(* Logix 5000 project; controller PLC_MCC1300_75F1 vendor 1 type 14 code 166 rev 32.11; software revision 32.04; part 9 of 83 *)

        [36].xFaulted := 1, [36].dEntryStatus := 16#0000_3000, [36].dFaultCode := 16#0000_0204, [36].dInstance := 16#0000_2268, [37].xConnected := 1, [37].xFaulted := 1, [37].dEntryStatus := 16#0000_3000, [37].dFaultCode := 16#0000_0204, [37].dInstance := 16#0000_494b, [38].xConnected := 1, [38].xFaulted := 1, [38].dEntryStatus := 16#0000_3000, [38].dFaultCode := 16#0000_0204, [38].dInstance := 16#0000_de82, [39].xConnected := 1, [39].xFaulted := 1, [39].dEntryStatus := 16#0000_3000, [39].dFaultCode := 16#0000_0204, [39].dInstance := 16#0000_ad3d, [40].xConnected := 1, [40].xFaulted := 1, [40].dEntryStatus := 16#0000_3000, [40].dFaultCode := 16#0000_0204, [40].dInstance := 16#0000_11ec, [41].xFaulted := 1, [41].dEntryStatus := 16#0000_1000, [41].dFaultCode := 16#0000_0204, [41].dInstance := 16#0000_7d3f, [42].xConnected := 1, [42].xFaulted := 1, [42].dEntryStatus := 16#0000_3000, [42].dFaultCode := 16#0000_0204, [42].dInstance := 16#0000_cb26, [43].xConnected := 1, [43].xFaulted := 1, [43].dEntryStatus := 16#0000_3000, [43].dFaultCode := 16#0000_0204, [43].dInstance := 16#0000_9dd1, [44].xConnected := 1, [44].xFaulted := 1, [44].dEntryStatus := 16#0000_3000, [44].dFaultCode := 16#0000_0204, [44].dInstance := 16#0000_2cb0, [45].xConnected := 1, [45].xFaulted := 1, [45].dEntryStatus := 16#0000_3000, [45].dFaultCode := 16#0000_0204, [45].dInstance := 16#0000_3773, [46].xConnected := 1, [46].xFaulted := 1, [46].dEntryStatus := 16#0000_3000, [46].dFaultCode := 16#0000_0204, [46].dInstance := 16#0000_0d0a, [47].xConnected := 1, [47].dEntryStatus := 16#0000_4000, [47].dInstance := 16#0000_f22b, [48].xConnected := 1, [48].dEntryStatus := 16#0000_4000, [48].dInstance := 16#0000_f6c7, [49].xConnected := 1,
        [49].dEntryStatus := 16#0000_4000, [49].dInstance := 16#0000_de7a); {access Read Only}
        [0]   // ETH_MCC1300
        [11]   // M3AZ01
        [12]   // M3AZ02
        [13]   // M3AZ03
        [14]   // M3AZ04
        [15]   // M3AZ05
        [16]   // M3AZ06
        [17]   // M3AZ07
        [18]   // M3AZ08
        [72]   // E93AZ1
        [31]   // TDKAZ05N
        [32]   // TDKAZ05S
        [33]   // TDAZ00N
        [34]   // TDAZ00S
        [35]   // TDAZ01N
        [36]   // TDAZ01S
        [37]   // TDAZ02N
        [19]   // M3AZ09
        [73]   // E96AZ1
        [75]   // E98AZ1
        [74]   // E97AZ1
        [20]   // M3AZ10
        [21]   // TDKAZ00N
        [38]   // TDAZ02S
        [39]   // TDAZ03N
        [40]   // TDAZ03S
        [41]   // TDAZ04N
        [42]   // TDAZ04S
        [43]   // TDAZ05N
        [44]   // TDAZ05S
        [50]   // E53AZ1
        [46]   // D010M1PM1
        [47]   // D010M2PM1
        [61]   // E77AZ1
        [62]   // E78AZ1
        [48]   // D020PM1
        [51]   // E61AZ1
        [52]   // E62AZ1
        [63]   // E81AZ1
        [64]   // E82AZ1
        [54]   // E64AZ1
        [53]   // E63AZ1
        [55]   // E65AZ1
        [65]   // E83AZ1
        [66]   // E84AZ1
        [56]   // E66AZ1
        [57]   // E67AZ1
        [58]   // E71AZ1
        [67]   // E85AZ1
        [68]   // E86AZ1
        [5]   // TD5680AP1
        [59]   // E73AZ1
        [60]   // E76AZ1
        [69]   // E87AZ1
        [70]   // E88AZ1
        [71]   // E91AZ1
        [1]   // ETH_M2
        [6]   // M3683AP1
        [7]   // E152AP1
        [8]   // RIOM13
        [22]   // TDKAZ00S
        [23]   // TDKAZ01N
        [24]   // TDKAZ01S
        [25]   // TDKAZ02N
        [26]   // TDKAZ02S
        [27]   // TDKAZ03N
        [28]   // TDKAZ03S
        [29]   // TDKAZ04N
        [30]   // TDKAZ04S
   MMI_DATA : INT[64] := ([1] := 4088, [2] := 4095, [8] := 4095, [11] := 2048, [20] := -1, [21] := -1, [22] := 1, [23] := 1);   // MMI DATA For Fix 32
        [12].0   // FIX MMI VMCC M2 Panel Overtemp Alarm
        [12].1   // FIX MMI VMCC TD Panel Overtemp Alarm
   MMI_FROM_MB : MESSAGE;
        MessageParameters(ServiceCode := 16#004b, LocalElement := MMI_DATA[20], ...)
   MMI_TO_MB : MESSAGE;
        MessageParameters(ServiceCode := 16#004c, LocalElement := MMI_DATA[0], ...)
   MMI_TO_MB_N15 : MESSAGE;
        MessageParameters(ServiceCode := 16#004c, LocalElement := MMI_DATA[0], ...)
   MS_LEHR : ALIAS FOR N20[11];
   MS_LINE : ALIAS FOR N20[13];
   MS_TRIM : ALIAS FOR N20[12];
   N10 : DINT[50] := ([10] := 2100, [40] := 4095);
        [16].1   // LEHR SPEED Speed received From Reliance Capping system is Valid
        [16].0   // LEHR SPEED Speed received From Reliance AutoMax PLC Is Valid
   N100 : DINT[1];
   N105 : DINT[1];
   N11 : DINT[500];
        [96]   // VISION INTERFACE: 2ND MOST CURRNET REJECTION REASON
        [97]   // VISION INTERFACE: 3RD MOST CURRNET REJECTION REASON
        [94].1   // Host & HMI Read Data: No Data From Vision System
        [94].2   // Host & HMI Read Data: Not Used Reserved for Focus CPS
        [94].3   // Host & HMI Read Data: Not Used Reserved for Focus CPS
        [94].4   // Host & HMI Read Data: Not Used Reserved for Focus CPS
        [79]   // Powder Camera Inspected Plate host IDENT
        [80]   // Host & HMI Read Data: Vision Broken Plate Count
        [81]   // Host & HMI Read Data: Vision Width Error Count
        [82]   // Host & HMI Read Data: Vision Length Error Count
        [83]   // Host & HMI Read Data: Vision Edge Defect Count
        [84]   // Host & HMI Read Data: Vision Corner Defect Count
        [85]   // Host & HMI Read Data: Vision Skew Count
        [86]   // Host & HMI Read Data: Vision Squareness Count
        [87]   // Host & HMI Read Data: Vision Fault Mark Count
        [88]   // Host & HMI Read Data: Vision Plate Missing Count
        [89]   // Host & HMI Read Data: Vision Not Separated Count
        [90]   // Host & HMI Read Data: Vision Other Count
        [91]   // Host & HMI Read Data: Vision Good Pieces Count
        [94].7   // Host & HMI Read Data: Vision System Is Disabled
        [92]   // Host & HMI Read Data: Vision Bad Pieces Count
        [93]   // Host & HMI Read Data: Vision No Response Count
        [94]   // Host & HMI Read Data: Vision Status Word
        [95]   // VISION INTERFACE: MOST CURRNET REJECTION REASON
        [94].0   // Host & HMI Read Data: All Pieces Are Bad
        [94].5   // Host & HMI Read Data: Vision System Is Online
        [94].6   // Host & HMI Read Data: Vision Service Required
   N110 : DINT[1];
   N115 : DINT[1];
   N11_HOST : INT[500] := ([0] := 22347, [1] := 22347, [20] := 9447, [21] := 96, [22] := 2047, [23] := 2047, [24] := 21845, [25] := 21, [26] := 53, [27] := 53, [38] := 2, [40] := 1, [60] := 554, [61] := 13, [62] := 20, [63] := 528, [65] := 609, [66] := 576, [67] := 4736, [68] := 453, [69] := 4902, [70] := 1028, [72] := 1536, [73] := 8320, [74] := 1, [79] := 8320, [80] := 1, [94] := 1, [101] := 648, [102] := 3, [103] := 204, [104] := 22347, [131] := 647, [133] := 45, [134] := 22346, [141] := 646, [143] := 45, [144] := 22346); {produced}
   N12 : DINT[500];
        [0]   // When this is Non-zero host Computer has Written new
        [3]   // HOST WRITE DATA: Glass Thickness (mils)
        [5]   // HOST WRITE DATA: Packing Station In Use Bits
        [6]   // HOST WRITE DATA: Ribbon Type (32=Eclipse Adv)
        [60]   // New cap data Buffer written by Host Computer
   N120 : DINT[1];
   N125 : DINT[1];
   N12_HOST : INT[500] := ([0] := 1, [1] := 650, [2] := 233, [3] := 15, [4] := 7653, [6] := 32, [7] := 31); {produced}
   N13 : DINT[500];
   N130 : INT[8] := ([0] := 1, [1] := 1, [2] := 1, [4] := 1325, [5] := 1, [6] := 1, [7] := 1);
        [3].10   // M2 -->> M4 Reliance Handoff Sensor (Redundant - on South side)
        [5].0   // M2-->M4 Benchboard No. 1 crusher Down
        [5].1   // M2-->M4 Benchboard No. 1 crusher Pushbutton
        [3].14   // M2 -->> M4 Crush all Selector Switch
        [3].15   // M2 -->> M4 Re-allocate To crusher Push-button
        [3].12   // M2 -->> M4 SPARE
        [3].1   // M2 -->> M4 SPARE
        [3].11   // M2 -->> M4
        [3].13   // M2 -->> M4 SPARE
        [3].2   // M2 -->> M4 SPARE
        [3].3   // M2 -->> M4 SPARE
        [3].4   // M2 -->> M4 SPARE
        [3].5   // M2 -->> M4 SPARE
        [3].6   // M2 -->> M4 SPARE
        [3].7   // M2 -->> M4 SPARE
        [3].8   // M2 -->> M4 SPARE
        [3].9   // M2 -->> M4 SPARE
   N131 : INT[8] := ([1] := 132, [4] := 450);
        [3].9   // M4 -->> M2 Reject Window Lamp
        [1]   // M2 -->> M4 Copy mainline Crusher status bits from M2 to M4
        [5].0   // M4-->M2 Float Glass Prodution
        [5].1   // M4-->M2 UL Crusher Is Faulted
        [3].14   // M4 -->> M2 ML is in Sleep Mode
        [3].3   // M4 -->> M2 Mainline Sec. Trans. Drive Fault
        [3].5   // M4 -->> M2 Mainline Sec. Trans. E-Stop
        [3].6   // M4 -->> M2 Mainline Sec. Trans. Backup
        [5].2   // M4-->M2 VISION SYS Rejected Plate Alarm Horn
        [1].11   // M4 -->> M2 Mainline vision Conveyor Stopped
        [3].10   // M4 -->> M2 Leg 2 Is In Sleep Mode Transfer Unavailable
        [3].11   // M4 -->> M2 Leg 3 Is In Sleep Mode Transfer Unavailable
        [3].12   // M4 -->> M2 Leg 4 Is In Sleep Mode Transfer Unavailable
        [3].13   // M4 -->> M2 Leg 5 Is In Sleep Mode Transfer Unavailable
        [4]   // M4 -->> M2 Trim speed
        [3].8   // M4 -->> M2 Reliance Data Received
        [3].15   // M4 -->> M2 M4 Heartbeat
        [3].1   // M4 -->> M2 SPARE
        [3].2   // M4 -->> M2 SPARE
   N135 : DINT[10];
        [0].12   // VHSC BTW Error Bit
        [5].12   // VHSC BTR Error Bit
        [0].15   // VHSC BTW Enable Bit
        [5].15   // VHSC BTR Enable Bit
   N136 : DINT[64];
        [1].15   // VHSC Data Representation Mode 0 = Binary 1 = BCD
        [30].0   // Output 01 Output/Counter Mapping Bits PC00
        [30].1   // Output 01 Output/Counter Mapping Bits PC01
        [30].2   // Output 01 Output/Counter Mapping Bits PC02
        [30].3   // Output 01 Output/Counter Mapping Bits PC03
        [1].0   // Reset PC00 - ACTIVE HIGH !
        [25].0   // Output 00 Output/Counter Mapping Bits PC00
        [25].1   // Output 00 Output/Counter Mapping Bits PC01
        [25].2   // Output 00 Output/Counter Mapping Bits PC02
        [25].3   // Output 00 Output/Counter Mapping Bits PC03
        [25]   // *************** * Output 00 ** * Mapping ** * Bits ** ***************
        [1].1   // Reset PC01 - ACTIVE HIGH !
        [21]   // Counter 0 Sample Period X 10mS
        [22]   // Counter 1 Sample Period X 10mS
        [1].2   // Reset PC02 - ACTIVE HIGH !
        [3]   // Mode Bits For Counters 0 and 1 ** Default ** ** Used **
        [13]   // PC00 Preset Value MSD
        [1].8   // PC00 Load Preset-
        [1].9   // PC01 Load Preset-
        [14]   // PC00 Preset Value LSD
        [15]   // PC01 Preset Value MSD
        [1].4   // PC00 New Data Acknowledge
        [2].10   // Output 02 Force
        [26]   // Output 00 ON VALUE MSD
        [10]   // PC02 Rollover Value LSD
        [11]   // PC03 Rollover Value LSD
        [12]   // PC03 Rollover Value LSD
        [16]   // PC01 Preset Value LSD
        [17]   // PC02 Preset Value MSD
        [18]   // PC02 Preset Value LSD
        [19]   // PC03 Preset Value LSD
        [1].10   // PC02 Load Preset-
        [1].11   // PC03 Load Preset-
        [5]   // PC00 Rollover Value MSD
        [1]   // Word 1 VHSC BTW Data
        [1].3   // Reset PC03 - ACTIVE HIGH !
        [6]   // PC00 Rollover Value LSD
        [7]   // PC01 Rollover Value MSD
        [1].12   // Not Used
        [1].13   // Not Used
        [1].14   // Not Used
        [1].5   // PC01 New Data Acknowledge
        [1].6   // PC03 New Data Acknowledge
        [1].7   // PC02 New Data Acknowledge
        [2].11   // Output 03 Force
        [2].12   // Output 04 Force
        [23]   // Counter 2 Sample Period X 10mS
        [24]   // Counter 3 Sample Period X 10mS
        [30]   // *************** * Output 01 ** * Mapping ** * Bits ** ***************
        [27]   // Output 00 ON VALUE LSD
        [31]   // Output 01 ON VALUE MSD
        [28]   // Output 00 OFF VALUE MSD
        [29]   // Output 00 OFF VALUE LSD
        [2]   // Word 2 VHSC BTW Data
        [2].0   // Output 00 Enable
        [2].1   // Output 01 Enable
        [2].13   // Output 05 Force
        [2].14   // Output 06 Force
        [2].15   // Output 07 Force
        [2].2   // Output 02 Enable
        [2].3   // Output 03 Enable
        [2].4   // Output 04 Enable
        [2].5   // Output 05 Enable
        [2].6   // Output 06 Enable
        [2].7   // Output 07 Enable
        [2].8   // Output 00 Force
        [2].9   // Output 01 Force
        [35]   // *************** * Output 02 ** * Mapping ** * Bits ** ***************
        [32]   // Output 01 ON VALUE LSD
        [36]   // Output 02 ON VALUE MSD
        [33]   // Output 01 OFF VALUE MSD
        [34]   // Output 01 OFF VALUE LSD
        [40]   // *************** * Output 03 ** * Mapping ** * Bits ** ***************
        [37]   // Output 02 ON VALUE LSD
        [46]   // Output 04 ON VALUE MSD
        [38]   // Output 02 OFF VALUE MSD
        [39]   // Output 02 OFF VALUE LSD
        [45]   // *************** * Output 04 ** * Mapping ** * Bits ** ***************
        [50]   // *************** * Output 05 ** * Mapping ** * Bits ** ***************
        [47]   // Output 04 ON VALUE LSD
        [56]   // Output 06 ON VALUE MSD
        [48]   // Output 04 OFF VALUE MSD
        [49]   // Output 04 OFF VALUE LSD
        [55]   // *************** * Output 06 ** * Mapping ** * Bits ** ***************
        [60]   // *************** * Output 07 ** * Mapping ** * Bits ** ***************
        [57]   // Output 06 ON VALUE LSD
        [61]   // Output 07 ON VALUE MSD
        [58]   // Output 06 OFF VALUE MSD
        [59]   // Output 06 OFF VALUE LSD
        [8]   // PC01 Rollover Value LSD
        [62]   // Output 07 ON VALUE LSD
        [63]   // Output 07 OFF VALUE MSD
        [9]   // PC02 Rollover Value MSD
   N137 : DINT[18];
   N138 : DINT[18];
   N139 : DINT[18];
        [1].0   // Successful First BTW after program start
        [2].10   // VHSC-PC02 Gate Input
        [1]   // VHSC status word No.1
        [1].10   // VHSC Gate Input
        [1].11   // VHSC Gate Input
        [2].8   // VHSC-PC00 Gate Input
        [10]   // PC03 Count LSD
        [2]   // VHSC status word No.2
        [1].8   // VHSC Gate Input
        [1].9   // VHSC Gate Input
        [2].0   // OUTPUT 00 Status
        [2].1   // OUTPUT 01 Status
        [2].12   // VHSC-PC03
        [2].13   // not used
        [2].15   // not used
        [2].2   // OUTPUT 02 Status
        [2].3   // OUTPUT 03 Status
        [2].4   // OUTPUT 04 Status
        [2].5   // OUTPUT 05 Status
        [2].6   // OUTPUT 06 Status
        [2].7   // OUTPUT 07 Status
        [2].9   // VHSC-PC01 Gate Input
        [3]   // PC00 Count MSD
        [4]   // PC00 Count LSD
        [5]   // PC01 Count MSD
        [6]   // PC01 Count LSD
        [7]   // PC02 Count MSD
        [8]   // PC02 Count LSD
        [9]   // PC03 Count LSD
   N14 : DINT[500] := ([61] := 4088, [62] := 4095, [68] := 4095, [71] := 2048, [80] := -1, [81] := -1, [82] := 1, [83] := 1, [240] := 6, [250] := 3313, [251] := 782, [260] := 7, [460] := 1, [469] := 258, [470] := 1, [479] := 258, [480] := -1, [488] := 256, [489] := 256, [490] := -1, [496] := 256, [497] := 256, [498] := 256, [499] := 256);
        [252].10   // TRIM DECK Trim Zone 5 North knocker Move Up
        [252].11   // TRIM DECK Trim Zone 5 South knocker Move Up
        [250].10   // TRIM DECK Trim Zone 5 North trim Auto mode
        [251].10   // TRIM DECK Trim Zone 5 North trim Manual mode
        [255]   // TRIM KNOCKERS Remapped inputs for all Move out Selector Sws.
        [273]   // TRIM DECK NTH Out Sel. Sw. Examine Masked Move Result
        [272]   // TRIM DECK NTH In Sel. Sw. Examine Masked Move Result
        [61]   // HOST/MMI READ Word containing Bits for drive Fault NORTH
        [253].10   // TRIM DECK Trim Zone 5 North knocker Move Down
        [240].1   // Float Glass Hold Down Wheels Manual Raise
        [256].0   // TRIM DECK Krurl drop North deck Move In
        [275]   // TRIM DECK STH In Sel. Sw. Examine Masked Move Result
        [253].2   // TRIM DECK Trim Zone 1 North knocker Move Down
        [276]   // TRIM DECK STH Out Sel. Sw. Examine Masked Move Result
        [251].11   // TRIM DECK Trim Zone 5 South trim Manual mode
        [253].3   // TRIM DECK Trim Zone 1 South knocker Move Down
        [256].1   // TRIM DECK Krurl drop South deck Move In
        [240].0   // Float Glass Hold Down Wheels Automatic Mode
        [250].2   // TRIM DECK Trim Zone 1 North trim Auto mode
        [260].0   // TRIM KNOCKERS Permissive to Start adj drive 1 = Drive idle 0 = Drv in use
        [255].10   // TRIM DECK Trim Zone 5 North knocker Move Out
        [255].11   // TRIM DECK Trim Zone 5 South knocker Move Out
        [271]   // TRIM DECK NTH Contactor Examine Masked Move Result
        [274]   // TRIM DECK STH Contactor Examine Masked Move Result
        [68]   // HOST/MMI READ Word containing Foward bits For Conveyors
        [253].4   // TRIM DECK Trim Zone 2 North knocker Move Down
        [253].5   // TRIM DECK Trim Zone 2 South knocker Move Down
        [253].6   // TRIM DECK Trim Zone 3 North knocker Move Down
        [253].7   // TRIM DECK Trim Zone 3 South knocker Move Down
        [254]   // TRIM KNOCKERS Remapped inputs for all Move in Selector Sws.
        [251].0   // TRIM DECK Krurl drop North trim Manual mode
        [460]   // TD MMI Zone 4 South Skew Adjustment
        [240].3   // Eclipse Hold Down Wheels Manual Raise
        [90].0   // To Float 1 host, bars on/off
        [312]   // HMI Data: Transfer 1A Stopping Offset for Rotated Glass [in x 10]
        [302]   // HMI Data: Transfer 1 Stopping Offset for Rotated Glass [in x 10]
        [351]   // HMI Read & Write Data: Transfer 1 Take All Cap Length
        [253].8   // TRIM DECK Trim Zone 4 North knocker Move Down
        [240].2   // Eclipse Hold Down Wheels Auto Mode
        [253].9   // TRIM DECK Trim Zone 4 South knocker Move Down
        [250].11   // TRIM DECK Trim Zone 5 South trim Auto mode
        [253].11   // TRIM DECK Trim Zone 5 South knocker Move Down
        [62]   // HOST/MMI READ Word containing Bits for drive Fault SOUTH AND 1-3
        [72].0   // FIX MMI VMCC M2 Panel Overtemp Alarm
        [72].1   // FIX MMI VMCC TD Panel Overtemp Alarm
        [470]   // TD MMI Zone 5 South Skew Adjustment
        [480]   // TD MMI Zone 3 South Skew Adjustment
        [490]   // TD MMI Zone 2 South Skew Adjustment
        [250]   // TRIM DECK Word containing All auto mode Bits
        [62].0   // Host Read Conv 1 Fault
        [251].2   // TRIM DECK Trim Zone 1 North trim Manual mode
        [250].3   // TRIM DECK Trim Zone 1 South trim Auto mode
        [61].10   // Host Read Conv 11N Fault
        [251].3   // TRIM DECK Trim Zone 1 South trim Manual mode
        [251].4   // TRIM DECK Trim Zone 2 North trim Manual mode
        [251].5   // TRIM DECK Trim Zone 2 South trim Manual mode
        [62].1   // Host Read Conv 2 Fault
        [61].11   // Host Read Conv 12N Fault
        [254].10   // TRIM DECK Trim Zone 5 North knocker Move In
        [254].11   // TRIM DECK Trim Zone 5 South knocker Move In
        [251].6   // TRIM DECK Trim Zone 3 North trim Manual mode
        [256].2   // TRIM DECK Trim Zone 1 North deck Move In
        [250].0   // TRIM DECK Krurl drop North trim Auto mode
        [250].4   // TRIM DECK Trim Zone 2 North trim Auto mode
        [256].3   // TRIM DECK Trim Zone 1 South deck Move In
        [251].7   // TRIM DECK Trim Zone 3 South trim Manual mode
        [251].8   // TRIM DECK Trim Zone 4 North trim Manual mode
        [256].4   // TRIM DECK Trim Zone 2 North deck Move In
        [251].9   // TRIM DECK Trim Zone 4 South trim Manual mode
        [256].5   // TRIM DECK Trim Zone 2 South deck Move In
        [250].1   // TRIM DECK Krurl drop South trim Auto mode
        [250].5   // TRIM DECK Trim Zone 2 South trim Auto mode
        [256].6   // TRIM DECK Trim Zone 3 North deck Move In
        [253].0   // TRIM DECK Krurl drop North knocker Move Down
        [253].1   // TRIM DECK Krurl drop South knocker Move Down
        [255].2   // TRIM DECK Trim Zone 1 North knocker Move Out
        [255].3   // TRIM DECK Trim Zone 1 South knocker Move Out
        [255].4   // TRIM DECK Trim Zone 2 North knocker Move Out
        [255].5   // TRIM DECK Trim Zone 2 South knocker Move Out
        [255].6   // TRIM DECK Trim Zone 3 North knocker Move Out
        [255].7   // TRIM DECK Trim Zone 3 South knocker Move Out
        [255].8   // TRIM DECK Trim Zone 4 North knocker Move Out
        [255].9   // TRIM DECK Trim Zone 4 South knocker Move Out
        [257].2   // TRIM DECK Trim Zone 1 North deck Move Out
        [256].7   // TRIM DECK Trim Zone 3 South deck Move In
        [257].3   // TRIM DECK Trim Zone 1 South deck Move Out
        [256].8   // TRIM DECK Trim Zone 4 North deck Move In
        [250].6   // TRIM DECK Trim Zone 3 North trim Auto mode
        [250].7   // TRIM DECK Trim Zone 3 South trim Auto mode
        [250].8   // TRIM DECK Trim Zone 4 North trim Auto mode
        [256].9   // TRIM DECK Trim Zone 4 South deck Move In
        [257].0   // TRIM DECK Krurl drop North deck Move Out
        [251].1   // TRIM DECK Krurl drop South trim Manual mode
        [252].2   // TRIM DECK Trim Zone 1 North knocker Move Up
        [257].4   // TRIM DECK Trim Zone 2 North deck Move Out
        [252].3   // TRIM DECK Trim Zone 1 South knocker Move Up
        [252].4   // TRIM DECK Trim Zone 2 North knocker Move Up
        [252].5   // TRIM DECK Trim Zone 2 South knocker Move Up
        [252].6   // TRIM DECK Trim Zone 3 North knocker Move Up
        [252].7   // TRIM DECK Trim Zone 3 South knocker Move Up
        [250].9   // TRIM DECK Trim Zone 4 South trim Auto mode
        [252].0   // TRIM DECK Krurl drop North knocker Move Up
        [252].1   // TRIM DECK Krurl drop South knocker Move Up
        [254].0   // TRIM DECK Krurl drop North knocker Move In
        [254].1   // TRIM DECK Krurl drop South knocker Move In
        [256].10   // TRIM DECK Trim Zone 5 North deck Move In
        [256].11   // TRIM DECK Trim Zone 5 South deck Move In
        [252].8   // TRIM DECK Trim Zone 4 North knocker Move Up
        [252].9   // TRIM DECK Trim Zone 4 South knocker Move Up
        [254].2   // TRIM DECK Trim Zone 1 North knocker Move In
        [254].3   // TRIM DECK Trim Zone 1 South knocker Move In
        [254].4   // TRIM DECK Trim Zone 2 North knocker Move In
        [254].5   // TRIM DECK Trim Zone 2 South knocker Move In
        [254].6   // TRIM DECK Trim Zone 3 North knocker Move In
        [254].7   // TRIM DECK Trim Zone 3 South knocker Move In
        [254].8   // TRIM DECK Trim Zone 4 North knocker Move In
        [254].9   // TRIM DECK Trim Zone 4 South knocker Move In
        [255].0   // TRIM DECK Krurl drop North knocker Move Out
        [255].1   // TRIM DECK Krurl drop South knocker Move Out
        [257].10   // TRIM DECK Trim Zone 5 North deck Move Out
        [257].11   // TRIM DECK Trim Zone 5 South deck Move Out
        [257].1   // TRIM DECK Krurl drop South deck Move Out
        [62].2   // Host Read Conv 3 Fault
        [84]   // HMI Write Data: Vision Edge On Defect Tol. [mm x 10]
        [112]   // HMI Write Data: Vision -Skew Tolerance [deg x 100]
        [80]   // HMI Write Data: Vision Over Width Tolerance [mm x 10]
        [301]   // HMI Data: Transfer 1 TE Stopping Position [in x 10]
        [257].5   // TRIM DECK Trim Zone 2 South deck Move Out
        [61].9   // Host Read Conv 10N Fault
        [62].9   // Host Read Conv 10S Fault
        [61].3   // Host Read Conv 4N Fault
        [257].6   // TRIM DECK Trim Zone 3 North deck Move Out
        [81]   // HMI Write Data: Vision Over Length Tolerance [mm x 10]
        [85]   // HMI Write Data: Vision Corner On Defect Tol. [mm x 10]
        [311]   // HMI Data: Transfer 1A TE Stopping Position [in x 10]
        [257].7   // TRIM DECK Trim Zone 3 South deck Move Out
        [110]   // HMI Write Data: Vision Under Width Tolerance [mm x 10]
        [111]   // HMI Write Data: Vision Under Length Tolerance [mm x 10]
        [114]   // HMI Write Data: Vision Edge Off Defect Tol. [mm x 10]
        [115]   // HMI Write Data: Vision Corner Off Defect Tol. [mm x 10]
        [170]   // MMI 400 DECK OP Adjust Distance For Larger Plates [in]
        [257].8   // TRIM DECK Trim Zone 4 North deck Move Out
        [250].12   // TRIM DECK SPARE
        [250].13   // TRIM DECK SPARE
        [250].14   // TRIM DECK SPARE
        [250].15   // TRIM DECK SPARE
        [251].12   // TRIM DECK SPARE
        [251].13   // TRIM DECK SPARE
        [251].14   // TRIM DECK SPARE
        [251].15   // TRIM DECK SPARE
        [252].12   // TRIM DECK SPARE
        [252].13   // TRIM DECK SPARE
        [252].14   // TRIM DECK SPARE
        [252].15   // TRIM DECK SPARE
        [253].12   // TRIM DECK SPARE
        [253].13   // TRIM DECK SPARE
        [253].14   // TRIM DECK SPARE
        [253].15   // TRIM DECK SPARE
        [254].12   // TRIM DECK SPARE
        [254].13   // TRIM DECK SPARE
        [254].14   // TRIM DECK SPARE
        [254].15   // TRIM DECK SPARE
        [255].12   // TRIM DECK SPARE
        [255].13   // TRIM DECK SPARE
        [255].14   // TRIM DECK SPARE
        [255].15   // TRIM DECK SPARE
        [256].12   // TRIM DECK SPARE
        [256].13   // TRIM DECK SPARE
        [256].14   // TRIM DECK SPARE
        [256].15   // TRIM DECK SPARE
        [257].12   // TRIM DECK SPARE
        [257].13   // TRIM DECK SPARE
        [257].14   // TRIM DECK SPARE
        [257].15   // TRIM DECK SPARE
        [257].9   // TRIM DECK Trim Zone 4 South deck Move Out
        [260].1   // TRIM DECK NTH Permissive to Start adj drive 1 = Drive idle 0 = Drv in use
        [260].2   // TRIM DECK STH Permissive to Start adj drive 1 = Drive idle 0 = Drv in use
        [62].10   // Host Read Conv 11S Fault
        [62].11   // Host Read Conv 12S Fault
        [61].4   // Host Read Conv 5N Fault
        [61].5   // Host Read Conv 6N Fault
        [61].6   // Host Read Conv 7N Fault
        [61].7   // Host Read Conv 8N Fault
        [61].8   // Host Read Conv 9N Fault
        [62].3   // Host Read Conv 4S Fault
        [62].4   // Host Read Conv 5S Fault
        [62].5   // Host Read Conv 6S Fault
        [62].6   // Host Read Conv 7S Fault
        [62].7   // Host Read Conv 8S Fault
        [62].8   // Host Read Conv 9S Fault
        [113]   // HMI Write Data: Vision -Squareness Tol. [mm x 10]
        [350]   // HMI Read & Write Data: Transfer 1 Take All Cap ID
        [358]   // HMI Read & Write Data: Transfer 1 Size A Split Width
        [82]   // HMI Write Data: Vision +Skew Tolerance [deg x 100]
        [83]   // HMI Write Data: Vision +Squareness Tol. [mm x 10]
        [86]   // HMI Write Data: Glass Substrate Type
   N14_HOST : INT[999]; {produced}
   N15 : DINT[500];
   N16 : DINT[500];
   N17 : DINT[100];
   N177 : DINT[10] := ([0] := 56, [1] := 1, [2] := 80, [5] := 2);
   N178 : DINT[100];
   N179 : DINT[100];
   N18 : DINT[100];
   N184 : DINT[50] := ([0] := 13, [1] := 94, [2] := 95, [3] := 96, [4] := 97, [5] := 98, [6] := 99, [7] := 100, [8] := 101, [9] := 4096, [10] := 11, [11] := 911, [12] := 671, [14] := 695, [16] := 23, [17] := 47, [18] := 107, [20] := 4, [21] := 139, [22] := 140, [23] := 141, [24] := 142, [25] := 143, [26] := 144, [27] := 145, [28] := 146, [29] := 8, [30] := 2, [31] := 902, [32] := 798, [34] := 686, [37] := 109, [49] := 2048);
   N185 : DINT[1];
   N187 : DINT[1];
   N188 : DINT[48] := ([4] := 256, [6] := 3840, [8] := 1280, [10] := 1280, [12] := 1280, [14] := 1280, [16] := 1280, [18] := 1280, [20] := 3328, [22] := 3840, [24] := 3840, [26] := 3840, [28] := 3840, [30] := 256);
   N189 : DINT[40];
   N190 : DINT[40];
   N191 : DINT[64];
   N192 : DINT[40];
   N193 : DINT[40] := ([0] := -22773, [1] := -27996, [5] := 1, [6] := 98, [7] := 1, [8] := 1, [17] := 102, [18] := 1, [20] := 96, [21] := 96, [22] := 97, [23] := 96, [24] := 97, [25] := 6, [26] := 103, [27] := 98, [28] := 98, [29] := 99, [30] := 474, [31] := 393, [32] := 96, [33] := 380);
   N194 : DINT[45] := ([2] := 166, [3] := 419, [4] := 166, [5] := 213, [7] := 206, [14] := -26651, [15] := 25346, [16] := 18332, [17] := -17337, [18] := 424, [19] := 19629, [20] := 169, [21] := 13674, [27] := 8, [29] := 1, [37] := 8114, [39] := 11259, [41] := 5595);
   N195 : DINT[40] := ([0] := 26204, [1] := 26204, [5] := 3, [7] := 1);
   N196 : DINT[1];
   N197 : DINT[1];
   N198 : DINT[1];
   N199 : DINT[1];
   N20 : DINT[50] := ([1] := 200, [2] := 500, [3] := 1200, [4] := 3000, [11] := 600, [12] := 150, [13] := 67, [14] := 40);
        [12]   // Milliseconds for two inches of glass travel at TRIM SPEED
        [11]   // Milliseconds for 2 inches of glass travel at LEHR SPEED
        [13]   // Milliseconds for 2 inches of glass travel at LINE SPEED
        [4]   // Runout Speed
        [1]   // Lehr Speed
        [2]   // Trim Speed
        [3]   // Line-Speed
   N200 : DINT[160];
   N201 : DINT[100];
   N202 : DINT[100];
   N203 : DINT[100];
   N204 : DINT[100];
   N205 : DINT[100];
   N206 : DINT[100];
   N207 : DINT[100];
   N208 : DINT[100];
   N209 : DINT[100];
   N21 : DINT[31] := ([0] := 2, [1] := 6144, [2] := 8320, [14] := 128);
        [0].5   // PLC -->> Copro Force Baseline/ Threshold (Set by MMI and Reset on LE)
        [0].2   // PLC -->> Copro Send Test Message to Vision
        [0].8   // PLC -->> Copro Reset Request for Baseline (Pushbutton at Vision)
        [0].3   // PLC -->> Copro No Update (From MMI)
        [14].8   // Copro -->> PLC Sending Test Message
        [14].0   // Copro -->> PLC All Bad Msg From Vision (Flashing Red)
        [14].1   // Copro -->> PLC No Data Msg From Vision (Solid Red)
        [0].1   // New data is Ready for VISCOMM Cleared by MLVISION
        [3]   // VISCOM Result Register --------------- 1=Good! 2=BAD!
        [0].4   // PLC --> Copro Reset Vision Counters (From VAX)
        [14].4   // Copro -->> PLC Doing Baseline (Flashing Blue)
        [14].5   // Copro -->> PLC Doing Threshold (Flasing Blue)
        [3].1   // VISCOM Result Register --------------- 1=Good! 2=Bad!
        [14].7   // Copro -->> PLC Copro Request for Baseline (Solid Blue)
        [3].0   // VISCOM Result Register --------------- 1 = Good 2 = Bad!
        [0].14   // PLC -->> Copro Used by VISCOM
        [14].6   // Copro -->> PLC Waiting
        [14].14   // Copro -->> PLC Bad Checksum
        [14].15   // Copro -->> PLC Bad Response
        [1]   // VISCOM New Length data (64ths)
        [2]   // VISCOM New Width data (64ths)
        [0].0   // PLC -->> Copro Debug
   N210 : DINT[100];
   N211 : DINT[100];
   N212 : DINT[100];
   N213 : DINT[100];
   N214 : DINT[100];
   N214_1 : ALIAS FOR N214[1];
   N214_5 : ALIAS FOR N214[5];
   N215 : DINT[100];
   N216 : DINT[100];
   N217 : DINT[100];
   N218 : DINT[100];
   N219 : DINT[100];
   N220 : DINT[100];
   N221 : DINT[100];
   N222 : DINT[100];
   N223 : DINT[100];
   N224 : DINT[100];
   N225 : DINT[100];
   N226 : DINT[100];
   N227 : DINT[100];
   N228 : DINT[100];
   N229 : DINT[100];
   N230 : DINT[100];
   N231 : DINT[100];
   N232 : DINT[100];
   N25 : DINT[110] := ([0] := 774, [1] := 1, [2] := 1, [3] := 1, [4] := 1, [5] := 1, [100] := 774);
        [1].1   // Vision System Results Buffer: Service Required for Vision System
        [3]   // Vision System Results Buffer: Number of Streams across Conveyor
        [0]   // Vision System Results Buffer: Group ID
        [2]   // Vision System Results Buffer: New data Flag (1 = New data)
        [100]   // Vision System Results PLC ID DTR Change of Value Reference
        [10]   // Vision System Results Buffer: Split 2B Reject Flag
        [11]   // Vision System Results Buffer: Split 2C Reject Flag
        [12]   // Vision System Results Buffer: Split 2D Reject Flag
        [13]   // Vision System Results Buffer: Split 3A Reject Flag
        [14]   // Vision System Results Buffer: Split 3B Reject Flag
        [15]   // Vision System Results Buffer: Split 3C Reject Flag
        [16]   // Vision System Results Buffer: Split 3D Reject Flag
        [17]   // Vision System Results Buffer: Split 4A Reject Flag
        [18]   // Vision System Results Buffer: Split 4B Reject Flag
        [19]   // Vision System Results Buffer: Split 4C Reject Flag
        [20]   // Vision System Results Buffer: Split 4D Reject Flag
        [21]   // Vision System Results Buffer: Split 5A Reject Flag
        [22]   // Vision System Results Buffer: Split 5B Reject Flag
        [23]   // Vision System Results Buffer: Split 5C Reject Flag
        [24]   // Vision System Results Buffer: Split 5D Reject Flag
        [25]   // Vision System Results Buffer: Split 6A Reject Flag
        [5]   // Vision System Results Buffer: Split 1A Reject Flag
        [6]   // Vision System Results Buffer: Split 1B Reject Flag
        [7]   // Vision System Results Buffer: Split 1C Reject Flag
        [26]   // Vision System Results Buffer: Split 6B Reject Flag
        [27]   // Vision System Results Buffer: Split 6C Reject Flag
        [28]   // Vision System Results Buffer: Split 6D Reject Flag
        [29]   // Vision System Results Buffer: Split 7A Reject Flag
        [30]   // Vision System Results Buffer: Split 7B Reject Flag
        [31]   // Vision System Results Buffer: Split 7C Reject Flag
        [32]   // Vision System Results Buffer: Split 7D Reject Flag
        [33]   // Vision System Results Buffer: Split 8A Reject Flag
        [34]   // Vision System Results Buffer: Split 8B Reject Flag
        [35]   // Vision System Results Buffer: Split 8C Reject Flag
        [36]   // Vision System Results Buffer: Split 8D Reject Flag
        [37]   // Vision System Results Buffer: Split 9A Reject Flag
        [38]   // Vision System Results Buffer: Split 9B Reject Flag
        [39]   // Vision System Results Buffer: Split 9C Reject Flag
        [40]   // Vision System Results Buffer: Split 9D Reject Flag
        [8]   // Vision System Results Buffer: Split 1D Reject Flag
        [9]   // Vision System Results Buffer: Split 2A Reject Flag
        [1]   // Vision System Results Buffer: Eagle-I Status Word
        [1].0   // Vision System Results Buffer: Vision System is Online
        [4]   // Vision System Results Buffer: Number of Splits down Conveyor
   N26 : DINT[150] := ([0] := 774, [2] := 3123, [3] := 1, [4] := 1, [5] := 12, [6] := 12, [7] := 1500, [8] := 32, [9] := 24, [10] := 32, [11] := 12, [12] := 12, [13] := 1500, [14] := 32, [15] := 24, [16] := 56, [17] := 8320, [21] := 5062, [100] := 20480, [101] := 774, [102] := 512, [105] := -22762, [106] := 2378, [107] := 23012, [108] := 4404, [109] := 22405, [110] := 846, [111] := -32768);
        [100].10   // VISION INTFCE: Cap Detected Entering Vision is a GOOD Plate with NO Splits
        [100].12   // VISION INTERFACE: Ignore Length Measurements on Queued Plates
        [100].2   // VISION INTERFACE: Results for New Cap ID Are Detected
        [100].4   // VISION INTERFACE: Cap Entering Conv 14 Check for Vis Required
        [100].8   // VIS INTFCE: Inspected Cap Prim Destination is Leg 1 or Leg 1A or L3
        [102].2   // one shot for Leading Edge of Data Valid Signal from Vision Sys
        [102].3   // VISION INTFCE: Bit to Reset Vision Debug Counters (Manually set)
        [102].8   // One shot for Glass Type Changing to Eclipse Advantage
        [104].0   // VIS INTFCE: No Vis Results Received for Glass Passing Thru X1 toward 1A
        [104].1   // VIS INTFCE: Inspection Results Not Received AND Glass is being Thrown Away
        [105]   // VISION INTERFACE: DEBUG COUNTER # of Good Plates from Data Packet
        [106]   // VISION INTERFACE: DEBUG COUNTER # of Bad Plates from Data Packet
        [107]   // VISION INTERFACE: DEBUG COUNTER # of Uninspected Plates from Data
        [109]   // VISION INTERFACE: DEBUG COUNTER # of Bad Plates from I/O Signals
        [13]   // Vision System Input Datafile: Neg Skew Tolerance [deg x 100]
        [100].9   // VIS INTFCE: Inspected Cap is a Leg 2 ; 4; or 5 Cap
        [100].3   // VISION INTERFACE: OK to Use New Vision Results
        [102].9   // One shot for Glass Type Changing to Base Glass
        [17]   // Vision System Input Datafile: Stream A Width [64ths]
        [18]   // Vision System Input Datafile: Stream B Width [64ths]
        [19]   // Vision System Input Datafile: Stream C Width [64ths]
        [20]   // Vision System Input Datafile: Stream D Width [64ths]
        [21]   // Vision System Input Datafile: Split 1 Length [64ths]
        [22]   // Vision System Input Datafile: Split 2 Length [64ths]
        [30].0   // Vision System Input Datafile: Stream A Inspect bit for Split 1
        [30].1   // Vision System Input Datafile: Stream A Inspect bit for Split 2
        [30].2   // Vision System Input Datafile: Stream A Inspect bit for Split 3
        [30].3   // Vision System Input Datafile: Stream A Inspect bit for Split 4
        [30].4   // Vision System Input Datafile: Stream A Inspect bit for Split 5
        [30].5   // Vision System Input Datafile: Stream A Inspect bit for Split 6
        [30].6   // Vision System Input Datafile: Stream A Inspect bit for Split 7
        [30].7   // Vision System Input Datafile: Stream A Inspect bit for Split 8
        [30].8   // Vision System Input Datafile: Stream A Inspect bit for Split 9
        [31].0   // Vision System Input Datafile: Stream B Inspect bit for Split 1
        [31].1   // Vision System Input Datafile: Stream B Inspect bit for Split 2
        [31].2   // Vision System Input Datafile: Stream B Inspect bit for Split 3
        [31].3   // Vision System Input Datafile: Stream B Inspect bit for Split 4
        [31].4   // Vision System Input Datafile: Stream B Inspect bit for Split 5
        [31].5   // Vision System Input Datafile: Stream B Inspect bit for Split 6
        [31].6   // Vision System Input Datafile: Stream B Inspect bit for Split 7
        [31].7   // Vision System Input Datafile: Stream B Inspect bit for Split 8
        [31].8   // Vision System Input Datafile: Stream B Inspect bit for Split 9
        [32].0   // Vision System Input Datafile: Stream C Inspect bit for Split 1
        [32].1   // Vision System Input Datafile: Stream C Inspect bit for Split 2
        [32].2   // Vision System Input Datafile: Stream C Inspect bit for Split 3
        [32].3   // Vision System Input Datafile: Stream C Inspect bit for Split 4
        [32].4   // Vision System Input Datafile: Stream C Inspect bit for Split 5
        [32].5   // Vision System Input Datafile: Stream C Inspect bit for Split 6
        [32].6   // Vision System Input Datafile: Stream C Inspect bit for Split 7
        [32].7   // Vision System Input Datafile: Stream C Inspect bit for Split 8
        [32].8   // Vision System Input Datafile: Stream C Inspect bit for Split 9
        [33].0   // Vision System Input Datafile: Stream D Inspect bit for Split 1
        [33].1   // Vision System Input Datafile: Stream D Inspect bit for Split 2
        [33].2   // Vision System Input Datafile: Stream D Inspect bit for Split 3
        [33].3   // Vision System Input Datafile: Stream D Inspect bit for Split 4
        [33].4   // Vision System Input Datafile: Stream D Inspect bit for Split 5
        [33].5   // Vision System Input Datafile: Stream D Inspect bit for Split 6
        [33].6   // Vision System Input Datafile: Stream D Inspect bit for Split 7
        [33].7   // Vision System Input Datafile: Stream D Inspect bit for Split 8
        [33].8   // Vision System Input Datafile: Stream D Inspect bit for Split 9
        [100].7   // VISION INTERFACE: Piece Called Bad By Vision Sys
        [102].10   // One shot for Glass Type Changing to Mirrorpane
        [34]   // Vision System Input Datafile: Quality Code for Split 1
        [35]   // Vision System Input Datafile: Quality Code for Split 2
        [36]   // Vision System Input Datafile: Quality Code for Split 3
        [37]   // Vision System Input Datafile: Quality Code for Split 4
        [38]   // Vision System Input Datafile: Quality Code for Split 5
        [39]   // Vision System Input Datafile: Quality Code for Split 6
        [40]   // Vision System Input Datafile: Quality Code for Split 7
        [15]   // Vision System Input Datafile: Neg Edge Tolerance [64ths]
        [6]   // Vision System Input Datafile: Pos Length Tolerance [64ths]
        [41]   // Vision System Input Datafile: Quality Code for Split 8
        [8]   // Vision System Input Datafile: Pos Square Tolerance [64ths]
        [99].0   // VISION INTERFACE: Primary Dest Cap Entering: Leg 1AN
        [99].1   // VISION INTERFACE: Primary Dest Cap Entering: Leg 1AS
        [99].2   // VISION INTERFACE: Primary Dest Cap Entering: Leg 1BN
        [99].4   // VISION INTERFACE: Primary Dest Cap Entering: Leg 2A LES
        [3]   // Vision System Input Datafile: Number of Streams across Conveyor
        [99].5   // VISION INTERFACE: Primary Dest Cap Entering: Leg 2B Robot
        [42]   // Vision System Input Datafile: Quality Code for Split 9
        [99]   // VISION INTERFACE: Primary Dest Cap Entering Vision Sys
        [1]   // Vision System Input Datafile: Substrate Type
        [100].5   // VISION INTERFACE: Cap Needs Vision Res Check for Receipt
        [100].0   // VISION INTERFACE: Cap Detected Entering the Vision System
        [23]   // Vision System Input Datafile: Split 3 Length [64ths]
        [24]   // Vision System Input Datafile: Split 4 Length [64ths]
        [9]   // Vision System Input Datafile: Pos Edge Tolerance [64ths]
        [11]   // Vision System Input Datafile: Neg Width Tolerance [64ths]
        [25]   // Vision System Input Datafile: Split 5 Length [64ths]
        [99].6   // VISION INTERFACE: Primary Dest Cap Entering: Mainline LES
        [99].3   // VISION INTERFACE: Primary Dest Cap Entering: Leg 1BS
        [100].15   // VISION INTERFACE: is Mirrorpane
        [0]   // Vision System Input Datafile: Group ID
        [101]   // VISION INTERFACE: PLC ID of Cap Entering Vision Sys
        [100].14   // VISION INTERFACE: Glass Type is Base glass
        [102].1   // One Shot for Glass Entering Conveyor 14
        [104].2   // VISION INTERFACE: Glass Type is Solar E
        [26]   // Vision System Input Datafile: Split 6 Length [64ths]
        [27]   // Vision System Input Datafile: Split 7 Length [64ths]
        [104].4   // VISION INTERFACE: Glass Type is TEC
        [28]   // Vision System Input Datafile: Split 8 Length [64ths]
        [29]   // Vision System Input Datafile: Split 9 Length [64ths]
        [104].5   // VISION INTERFACE: Glass Type is MirrorView
        [100].11   // VIS INTFCE: Glass Inspection Is in Progress
        [100].13   // VISION INTERFACE: Glass Type is Eclipse Adv
        [102].11   // One shot for Glass Type Changing to Solar E
        [103]   // VISION INTERFACE: Inspected Cap Primary Dest Word
        [30]   // Vision System Input Datafile: Stream A Inspect Word
        [31]   // Vision System Input Datafile: Stream B Inspect Word
        [32]   // Vision System Input Datafile: Stream C Inspect Word
        [33]   // Vision System Input Datafile: Stream D Inspect Word
        [100].6   // VISION INTERFACE: Piece Called Good By Vision Sys
        [102].12   // One shot for Glass Type Changing to Blue Active
        [2]   // Vision System Input Datafile: Substrate Thickness [64ths]
        [104].3   // VISION INTERFACE: Glass Type is Blue Active
        [102].0   // One Shot for Glass Entering Vision System
        [5]   // Vision System Input Datafile: Pos Width Tolerance [64ths]
        [100].1   // VISION INTERFACE: New Data Copied from Vision Output
        [10]   // Vision System Input Datafile: Pos Corner Tolerance [64ths]
        [12]   // Vision System Input Datafile: Neg Length Tolerance [64ths]
        [14]   // Vision System Input Datafile: Neg Square Tolerance [64ths]
        [16]   // Vision System Input Datafile: Neg Corner Tolerance [64ths]
        [4]   // Vision System Input Datafile: Number of Splits down Conveyor
        [7]   // Vision System Input Datafile: Pos Skew Tolerance [deg x 100]
        [108]   // VISION INTFCE: DEBUG COUNTER # of Good or Uninspected Plates from I/O signals
   N26_101 : ALIAS FOR N26[101];
   N27 : DINT[110] := ([0] := 774, [1] := 1, [3] := 1, [4] := 1, [5] := 1, [41] := 53, [42] := 52, [43] := 46, [44] := 54, [45] := 32, [46] := 32, [47] := 32, [48] := 82, [49] := 61, [50] := 48, [51] := 51, [52] := 55, [53] := 53, [54] := 53, [55] := 46, [56] := 53, [57] := 32, [58] := 32, [59] := 32, [60] := 1, [61] := 61, [62] := 48, [63] := 50, [64] := 49, [65] := 48, [66] := 53, [67] := 46, [68] := 48, [69] := 32, [70] := 32, [71] := 32, [72] := 87, [73] := 61, [74] := 48, [75] := 51, [76] := 51, [77] := 48, [78] := 48, [79] := 46, [80] := 57, [81] := 55, [82] := 13, [83] := 10);
        [1].1   // Vision System Results Buffer: Service Required for Vision System
        [3]   // Vision System Results Buffer: Number of Streams across Conveyor
        [0]   // Vision System Results Buffer: Group ID
        [2]   // Vision System Results Buffer: New data Flag (1 = New data)
        [10]   // Vision System Results Buffer: Split 2B Reject Flag
        [11]   // Vision System Results Buffer: Split 2C Reject Flag
        [12]   // Vision System Results Buffer: Split 2D Reject Flag
        [13]   // Vision System Results Buffer: Split 3A Reject Flag
        [14]   // Vision System Results Buffer: Split 3B Reject Flag
        [15]   // Vision System Results Buffer: Split 3C Reject Flag
        [16]   // Vision System Results Buffer: Split 3D Reject Flag
        [60].0   // VISION SYSTEM Status Indicators: Heartbeat Signal
        [5]   // Vision System Results Buffer: Split 1A Reject Flag
        [60].3   // VISION SYSTEM Status Indicators: PLC Read Error Occurred
        [6]   // Vision System Results Buffer: Split 1B Reject Flag
        [17]   // Vision System Results Buffer: Split 4A Reject Flag
        [18]   // Vision System Results Buffer: Split 4B Reject Flag
        [7]   // Vision System Results Buffer: Split 1C Reject Flag
        [19]   // Vision System Results Buffer: Split 4C Reject Flag
        [20]   // Vision System Results Buffer: Split 4D Reject Flag
        [21]   // Vision System Results Buffer: Split 5A Reject Flag
        [22]   // Vision System Results Buffer: Split 5B Reject Flag
        [23]   // Vision System Results Buffer: Split 5C Reject Flag
        [24]   // Vision System Results Buffer: Split 5D Reject Flag
        [25]   // Vision System Results Buffer: Split 6A Reject Flag
        [60].1   // VISION SYSTEM Status Indicators: System Stopped (0 = Running 1 = Stopped)
        [8]   // Vision System Results Buffer: Split 1D Reject Flag
        [26]   // Vision System Results Buffer: Split 6B Reject Flag
        [27]   // Vision System Results Buffer: Split 6C Reject Flag
        [28]   // Vision System Results Buffer: Split 6D Reject Flag
        [29]   // Vision System Results Buffer: Split 7A Reject Flag
        [30]   // Vision System Results Buffer: Split 7B Reject Flag
        [31]   // Vision System Results Buffer: Split 7C Reject Flag
        [32]   // Vision System Results Buffer: Split 7D Reject Flag
        [33]   // Vision System Results Buffer: Split 8A Reject Flag
        [34]   // Vision System Results Buffer: Split 8B Reject Flag
        [35]   // Vision System Results Buffer: Split 8C Reject Flag
        [36]   // Vision System Results Buffer: Split 8D Reject Flag
        [37]   // Vision System Results Buffer: Split 9A Reject Flag
        [38]   // Vision System Results Buffer: Split 9B Reject Flag
        [39]   // Vision System Results Buffer: Split 9C Reject Flag
        [40]   // Vision System Results Buffer: Split 9D Reject Flag
        [9]   // Vision System Results Buffer: Split 2A Reject Flag
        [60].2   // VISION SYSTEM Status Indicators: Outputs are OFF (0 = Outputs ON 1 = Outputs OFF)
        [1]   // Vision System Results Buffer: Eagle-I Status Word
        [1].0   // Vision System Results Buffer: Vision System is Online
        [4]   // Vision System Results Buffer: Number of Splits down Conveyor
        [60]   // VISION SYSTEM Status word From Eagle-I
   N30 : DINT[32] := ([1] := -2096895798, [2] := -2096895798);
        [10]   // Conveyor 10 Millisecond Accumulator Updated by STI File 18
        [11]   // Conveyor 11 Millisecond Accumulator Updated by STI File 18
        [12]   // Conveyor 12 Millisecond Accumulator Updated by STI File 18
        [13]   // Conveyor 13 Millisecond Accumulator Updated by STI File 18
        [14]   // Conveyor 14 Millisecond Accumulator Updated by STI File 18
        [15]   // Conveyor 15 Millisecond Accumulator Updated by STI File 18
        [1]   // Conveyor 1 Millisecond Accumulator Updated by STI File 18
        [2]   // Conveyor 2 Millisecond Accumulator Updated by STI File 18
        [3]   // Conveyor 3 Millisecond Accumulator Updated by STI File 18
        [4]   // Conveyor 4 Millisecond Accumulator Updated by STI File 18
        [5]   // Conveyor 5 Millisecond Accumulator Updated by STI File 18